DATA_BLOCK "DB_Scada_default"   // DB2112
{ S7_Optimized_Access := 'FALSE' }
VERSION : 0.1
   VAR
      tAlm : Struct   // HMI Alarms
         tE : Struct
            x0 : Bool;   // KE.Main emergency on
            x1 : Bool;   // KE1.Local emergency on
            x2 : Bool;   // Cabinet.Emergency localization
            x3 : Bool;   // SB1.Emergency localization
            x4 : Bool;   // SB2.Emergency localization
            x5 : Bool;
            x6 : Bool;
            x7 : Bool;
            x8 : Bool;
            x9 : Bool;
            x10 : Bool;
            x11 : Bool;
            x12 : Bool;
            x13 : Bool;
            x14 : Bool;
            x15 : Bool;
            x16 : Bool;
            x17 : Bool;
            x18 : Bool;
            x19 : Bool;
            x20 : Bool;
            x21 : Bool;
            x22 : Bool;
            x23 : Bool;
            x24 : Bool;
            x25 : Bool;
            x26 : Bool;
            x27 : Bool;
            x28 : Bool;
            x29 : Bool;
            x30 : Bool;
            x31 : Bool;
         END_STRUCT;
         tS : Struct
            tS0 : Struct
               x0 : Bool;
               x1 : Bool;   // Syncro.YCut meter gap outside the limits
               x2 : Bool;
               x3 : Bool;
               x4 : Bool;
               x5 : Bool;
               x6 : Bool;
               x7 : Bool;
               x8 : Bool;   // xB21QF1.Power supply 24V logic
               x9 : Bool;
               x10 : Bool;   // Syncro.Main line meter gap outside the limits
               x11 : Bool;
               x12 : Bool;
               x13 : Bool;
               x14 : Bool;
               x15 : Bool;
               x16 : Bool;
               x17 : Bool;
               x18 : Bool;
               x19 : Bool;
               x20 : Bool;
               x21 : Bool;
               x22 : Bool;
               x23 : Bool;
               x24 : Bool;
               x25 : Bool;
               x26 : Bool;
               x27 : Bool;
               x28 : Bool;
               x29 : Bool;
               x30 : Bool;
               x31 : Bool;
            END_STRUCT;
            tS1 : Struct
               x0 : Bool;
               x1 : Bool;   // Syncro.YCut meter gap outside the limits
               x2 : Bool;
               x3 : Bool;
               x4 : Bool;
               x5 : Bool;
               x6 : Bool;
               x7 : Bool;
               x8 : Bool;   // xB21QF1.Power supply 24V logic
               x9 : Bool;
               x10 : Bool;   // Syncro.Main line meter gap outside the limits
               x11 : Bool;
               x12 : Bool;
               x13 : Bool;
               x14 : Bool;
               x15 : Bool;
               x16 : Bool;
               x17 : Bool;
               x18 : Bool;
               x19 : Bool;
               x20 : Bool;
               x21 : Bool;
               x22 : Bool;
               x23 : Bool;
               x24 : Bool;
               x25 : Bool;
               x26 : Bool;
               x27 : Bool;
               x28 : Bool;
               x29 : Bool;
               x30 : Bool;
               x31 : Bool;
            END_STRUCT;
            tS2 : Struct
               x0 : Bool;
               x1 : Bool;   // Syncro.YCut meter gap outside the limits
               x2 : Bool;
               x3 : Bool;
               x4 : Bool;
               x5 : Bool;
               x6 : Bool;
               x7 : Bool;
               x8 : Bool;   // xB21QF1.Power supply 24V logic
               x9 : Bool;
               x10 : Bool;   // Syncro.Main line meter gap outside the limits
               x11 : Bool;
               x12 : Bool;
               x13 : Bool;
               x14 : Bool;
               x15 : Bool;
               x16 : Bool;
               x17 : Bool;
               x18 : Bool;
               x19 : Bool;
               x20 : Bool;
               x21 : Bool;
               x22 : Bool;
               x23 : Bool;
               x24 : Bool;
               x25 : Bool;
               x26 : Bool;
               x27 : Bool;
               x28 : Bool;
               x29 : Bool;
               x30 : Bool;
               x31 : Bool;
            END_STRUCT;
            tS3 : Struct
               x0 : Bool;
               x1 : Bool;   // Syncro.YCut meter gap outside the limits
               x2 : Bool;
               x3 : Bool;
               x4 : Bool;
               x5 : Bool;
               x6 : Bool;
               x7 : Bool;
               x8 : Bool;   // xB21QF1.Power supply 24V logic
               x9 : Bool;
               x10 : Bool;   // Syncro.Main line meter gap outside the limits
               x11 : Bool;
               x12 : Bool;
               x13 : Bool;
               x14 : Bool;
               x15 : Bool;
               x16 : Bool;
               x17 : Bool;
               x18 : Bool;
               x19 : Bool;
               x20 : Bool;
               x21 : Bool;
               x22 : Bool;
               x23 : Bool;
               x24 : Bool;
               x25 : Bool;
               x26 : Bool;
               x27 : Bool;
               x28 : Bool;
               x29 : Bool;
               x30 : Bool;
               x31 : Bool;
            END_STRUCT;
         END_STRUCT;
         tF : Struct
            x0 : Bool;
            x1 : Bool;
            x2 : Bool;
            x3 : Bool;
            x4 : Bool;
            x5 : Bool;
            x6 : Bool;
            x7 : Bool;
            x8 : Bool;
            x9 : Bool;
            x10 : Bool;
            x11 : Bool;
            x12 : Bool;
            x13 : Bool;
            x14 : Bool;
            x15 : Bool;
            x16 : Bool;
            x17 : Bool;
            x18 : Bool;
            x19 : Bool;
            x20 : Bool;
            x21 : Bool;
            x22 : Bool;
            x23 : Bool;
            x24 : Bool;
            x25 : Bool;
            x26 : Bool;
            x27 : Bool;
            x28 : Bool;
            x29 : Bool;
            x30 : Bool;
            x31 : Bool;
         END_STRUCT;
         tW : Struct
            x0 : Bool;   // PLCA.Timeout receiving consumed message
            x1 : Bool;   // PLCB.Timeout receiving consumed message
            x2 : Bool;   // PLCA.Mission packet lost
            x3 : Bool;   // PLCB.Mission packet lost
            x4 : Bool;   // PLCA.Syncro packet lost
            x5 : Bool;   // PLCB.Syncro packet lost
            x6 : Bool;   // QF.Protection air conditioners
            x7 : Bool;
            x8 : Bool;
            x9 : Bool;
            x10 : Bool;
            x11 : Bool;
            x12 : Bool;
            x13 : Bool;
            x14 : Bool;
            x15 : Bool;
            x16 : Bool;
            x17 : Bool;
            x18 : Bool;
            x19 : Bool;
            x20 : Bool;
            x21 : Bool;
            x22 : Bool;
            x23 : Bool;
            x24 : Bool;
            x25 : Bool;
            x26 : Bool;
            x27 : Bool;
            x28 : Bool;
            x29 : Bool;
            x30 : Bool;
            x31 : Bool;
         END_STRUCT;
      END_STRUCT;
      tHMR : Struct   // HMI Read
         xSpare0 : Bool := FALSE;   // Calibration function allowed {x|x|x|x|O}
         xSpare1 : Bool;
         xSpare2 : Bool;
         xSpare3 : Bool;
         xSpare4 : Bool;
         xSpare5 : Bool;
         xSpare6 : Bool;
         xSpare7 : Bool;
         xSpare8 : Bool;
         xSpare9 : Bool;
         xSpare10 : Bool;
         xSpare11 : Bool;
         xSpare12 : Bool;
         xSpare13 : Bool;
         xSpare14 : Bool;
         xSpare15 : Bool := FALSE;
         xSpare16 : Bool;
         xSpare17 : Bool;
         xSpare18 : Bool;
         xSpare19 : Bool;
         xSpare20 : Bool;
         xSpare21 : Bool;
         xSpare22 : Bool;
         xSpare23 : Bool;
         xSpare24 : Bool;
         xSpare25 : Bool;
         xSpare26 : Bool;
         xSpare27 : Bool;
         xSpare28 : Bool;
         xSpare29 : Bool;
         xSpare30 : Bool;
         xSpare31 : Bool;
         xSpare : Array[0..15] of Bool;
         iSpare0 : Int;
         iSpare1 : Int;
         iSpare2 : Int;
         iSpare3 : Int;
         iSpare4 : Int;
         iSpare5 : Int;
         iSpare6 : Int;
         iSpare7 : Int;
         iSpare8 : Int;
         iSpare9 : Int;
         iSpare10 : Int;
         iSpare11 : Int;
         iSpare12 : Int;
         iSpare13 : Int;
         iSpare14 : Int;
         iSpare15 : Int;
         iSpare16 : Int;
         dSpare0 : DInt := 0;   // Zone modality (1=Manual;4=Automatic;8=Manual request) {x|x|x|x|O}
         dSpare1 : DInt := 0;   // HMI Alarms
         dSpare2 : DInt := 0;   // HMI Write
         dSpare3 : DInt := 0;   // Production modality request (1=Out of Production 3= In production) {x|x|x|x|O}
         dSpare4 : DInt := 0;   // Production modality actual (1=Out of production 3=In production 8=Out of production request 9=In production request) {x|x|x|x|O}
         dSpare5 : DInt := 0;
         dSpare6 : DInt := 0;
         dSpare7 : DInt := 0;
         dSpare8 : DInt := 0;
         dSpare9 : DInt := 0;
         dSpare10 : DInt := 0;
         dSpare11 : DInt := 0;
         dSpare12 : DInt;
         dSpare13 : DInt;
         dSpare14 : DInt;
         dSpare15 : DInt;
         dSpare : Array[0..15] of DInt;
         rSpare0 : Real;
         rSpare1 : Real;
         rSpare2 : Real;
         rSpare3 : Real;
         rSpare4 : Real;
         rSpare5 : Real;
         rSpare6 : Real;
         rSpare7 : Real;
         rSpare8 : Real;
         tManCmd : Struct
            xSpare0 : Bool;
            xSpare1 : Bool;
            xSpare2 : Bool;
            xSpare3 : Bool;
            xSpare4 : Bool;
            xSpare5 : Bool;
            xSpare6 : Bool;
            xSpare7 : Bool;
            xSpare8 : Bool;
            xSpare9 : Bool;
            xSpare10 : Bool;
            xSpare11 : Bool;
            xSpare12 : Bool;
            xSpare13 : Bool;
            xSpare14 : Bool;
            xSpare15 : Bool;
            xSpare : Array[0..15] of Bool;
         END_STRUCT;
      END_STRUCT;
      tHMW : Struct   // HMI Write
         xSpare0 : Bool := FALSE;   // Automatic mode request {x|x|x|x|O}
         xSpare1 : Bool := FALSE;   // Manual mode request {x|x|x|x|O}
         xSpare2 : Bool := FALSE;   // Bridge out of production request {x|x|x|x|O}
         xSpare3 : Bool := FALSE;   // Bridge in production request {x|x|x|x|O}
         xSpare4 : Bool := FALSE;   // Cut during glass break {x|x|x|x|O}
         xSpare5 : Bool := FALSE;   // Motors and cards initialize {x|x|x|x|M}
         xSpare6 : Bool := FALSE;   // Force the homing of the heads {x|x|x|x|M}
         xSpare7 : Bool := FALSE;   // Position calibration request {x|x|x|x|M}
         xSpare8 : Bool := FALSE;   // Bridge offset calibration request {x|x|x|x|M}
         xSpare9 : Bool;
         xSpare10 : Bool;
         xSpare11 : Bool;
         xSpare12 : Bool;
         xSpare13 : Bool;
         xSpare14 : Bool := FALSE;
         xSpare15 : Bool := FALSE;
         xSpare16 : Bool := TRUE;
         xSpare17 : Bool := TRUE;
         xSpare18 : Bool := TRUE;
         xSpare19 : Bool := TRUE;
         xSpare20 : Bool := TRUE;
         xSpare21 : Bool := TRUE;
         xSpare22 : Bool := TRUE;
         xSpare23 : Bool := TRUE;
         xSpare24 : Bool;
         xSpare25 : Bool;
         xSpare26 : Bool;
         xSpare27 : Bool;
         xSpare28 : Bool;
         xSpare29 : Bool;
         xSpare30 : Bool;
         xSpare31 : Bool;
         xSpare : Array[0..15] of Bool;
         iSpare0 : Int;
         iSpare1 : Int;
         iSpare2 : Int;
         iSpare3 : Int;
         iSpare4 : Int;
         iSpare5 : Int;
         iSpare6 : Int;
         iSpare7 : Int;
         iSpare8 : Int;
         iSpare9 : Int;
         iSpare10 : Int;
         iSpare11 : Int;
         iSpare12 : Int;
         iSpare13 : Int;
         iSpare14 : Int;
         iSpare15 : Int;
         iSpare16 : Int := 0;
         dSpare0 : DInt := 0;   // Calibration. number of lite on calibration {x|x|1|8|M}
         dSpare1 : DInt := 0;   // Calibration. Move all the heads of this offset {mm/100|mm|-100|100|M}
         dSpare2 : DInt := 0;   // Pressure scaler during sample plate [%] {%|%|0|100|O}
         dSpare3 : DInt := 0;
         dSpare4 : DInt;
         dSpare5 : DInt;
         dSpare6 : DInt;
         dSpare7 : DInt;
         dSpare8 : DInt;
         dSpare9 : DInt;
         dSpare10 : DInt;
         dSpare11 : DInt;
         dSpare12 : DInt;
         dSpare13 : DInt;
         dSpare14 : DInt;
         dSpare15 : DInt;
         dSpare16 : DInt;
         dSpare17 : DInt;
         dSpare18 : DInt;
         dSpare19 : DInt;
         dSpare20 : DInt;
         dSpare21 : DInt;
         dSpare22 : DInt;
         dSpare23 : DInt;
         dSpare24 : DInt;
         dSpare25 : DInt;
         dSpare26 : DInt;
         dSpare27 : DInt;
         dSpare28 : DInt;
         dSpare29 : DInt;
         dSpare30 : DInt;
         dSpare31 : DInt;
         dSpare32 : DInt;
         dSpare33 : DInt;
         dSpare34 : DInt;
         dSpare35 : DInt;
         dSpare36 : DInt;
         dSpare37 : DInt;
         dSpare38 : DInt;
         dSpare39 : DInt;
         dSpare : Array[0..19] of DInt;
         rSpare0 : Real;
         rSpare1 : Real;
         rSpare2 : Real;
         rSpare3 : Real;
         rSpare4 : Real;
         rSpare5 : Real;
         rSpare6 : Real;
         rSpare7 : Real;
         rSpare8 : Real;
         tManCmd : Struct
            xSpare0 : Bool := FALSE;
            xSpare1 : Bool := FALSE;
            xSpare2 : Bool;
            xSpare3 : Bool;
            xSpare4 : Bool;
            xSpare5 : Bool;
            xSpare6 : Bool;
            xSpare7 : Bool;
            xSpare8 : Bool;
            xSpare9 : Bool;
            xSpare10 : Bool;
            xSpare11 : Bool;
            xSpare12 : Bool;
            xSpare13 : Bool;
            xSpare14 : Bool;
            xSpare15 : Bool;
            xSpare16 : Bool;
            xSpare17 : Bool;
            xSpare18 : Bool;
            xSpare19 : Bool;
            xSpare20 : Bool;
            xSpare21 : Bool;
            xSpare22 : Bool;
            xSpare23 : Bool;
            xSpare24 : Bool;
            xSpare25 : Bool;
            xSpare26 : Bool;
            xSpare27 : Bool;
            xSpare28 : Bool;
            xSpare29 : Bool;
            xSpare30 : Bool;
            xSpare31 : Bool;
         END_STRUCT;
      END_STRUCT;
   END_VAR
BEGIN
END_DATA_BLOCK

// folder: Communication

DATA_BLOCK "CM_Manager"   // DB1
{ S7_Optimized_Access := 'TRUE' }
VERSION : 0.1
BEGIN
END_DATA_BLOCK

DATA_BLOCK "CM_IDEV_FromMainLine"   // DB2
{ S7_Optimized_Access := 'TRUE' }
VERSION : 0.1
BEGIN
END_DATA_BLOCK

DATA_BLOCK "CM_IDEV_ToMainLine"   // DB3
{ S7_Optimized_Access := 'TRUE' }
VERSION : 0.1
BEGIN
END_DATA_BLOCK

DATA_BLOCK "CM_RECV_MissionData"   // DB4
{ S7_Optimized_Access := 'TRUE' }
VERSION : 0.1
BEGIN
END_DATA_BLOCK

DATA_BLOCK "CM_RECV_SyncroData"   // DB8
{ S7_Optimized_Access := 'TRUE' }
VERSION : 0.1
BEGIN
END_DATA_BLOCK

DATA_BLOCK "CM_BRCV_FromMainLine0"   // DB12
{ S7_Optimized_Access := 'TRUE' }
VERSION : 0.1
BEGIN
END_DATA_BLOCK

DATA_BLOCK "CM_BRCV_FromMainLine1"   // DB24
{ S7_Optimized_Access := 'TRUE' }
VERSION : 0.1
BEGIN
END_DATA_BLOCK

// folder: ILx2_Blocks

DATA_BLOCK "ILx2T_Parameter_Initialize_DB"   // DB10
{ S7_Optimized_Access := 'TRUE' }
VERSION : 1.1
// stored: InstanceOfName ILx2T_Parameter_Read_Write
"ILx2T_Parameter_Read_Write"
BEGIN
END_DATA_BLOCK

// folder: Subroutine

DATA_BLOCK "OB_Initialize"   // DB18
{ S7_Optimized_Access := 'TRUE' }
AUTHOR : Cigliutt
FAMILY : GP
VERSION : 1.0
// stored: InstanceOfName GP_OB_Initialize
"GP_OB_Initialize"
BEGIN
END_DATA_BLOCK

// folder: TaskErrors

DATA_BLOCK "RALRM_AUX_DB"   // DB59
{ S7_Optimized_Access := 'TRUE' }
VERSION : 0.1
   VAR RETAIN
      tAlm : Struct   // HMI Alarms
         tS : Struct   // Stopping faults
            xSpare_0 : Bool := FALSE;
            xSpare_1 : Bool := FALSE;
            xSpare_2 : Bool := FALSE;
            xSpare_3 : Bool := FALSE;
            xSpare_4 : Bool := FALSE;
            xSpare_5 : Bool := FALSE;
            xSpare_6 : Bool := FALSE;
            xSpare_7 : Bool := FALSE;
            xSpare_8 : Bool := FALSE;
            xSpare_9 : Bool := FALSE;
            xSpare_10 : Bool := FALSE;
            xSpare_11 : Bool := FALSE;
            xSpare_12 : Bool := FALSE;
            xSpare_13 : Bool := FALSE;
            xSpare_14 : Bool := FALSE;
            xSpare_15 : Bool := FALSE;
            xSpare_16 : Bool := FALSE;
            xSpare_17 : Bool := FALSE;
            xSpare_18 : Bool := FALSE;
            xSpare_19 : Bool := FALSE;
            xSpare_20 : Bool := FALSE;
            xSpare_21 : Bool := FALSE;
            xSpare_22 : Bool := FALSE;
            xSpare_23 : Bool := FALSE;
            xSpare_24 : Bool := FALSE;
            xSpare_25 : Bool := FALSE;
            xSpare_26 : Bool := FALSE;
            xSpare_27 : Bool := FALSE;
            xSpare_28 : Bool := FALSE;
            xSpare_29 : Bool := FALSE;
            xSpare_30 : Bool := FALSE;
            xSpare_31 : Bool := FALSE;
         END_STRUCT;
         tF : Struct   // Faults
            xDevice1 : Bool := FALSE;   // R13QF1.R13QF2.Power failure 230v auxiliary / Status device error.Device#1
            xDevice2 : Bool := FALSE;   // R18QF3.Power supply 24v logic / Status device error.Device#2
            xDevice3 : Bool := FALSE;   // R18QF4.Power supply 24v logic / Status device error.Device#3
            xDevice4 : Bool := FALSE;   // R18AP1.Redundancy 24v ok / Status device error.Device#4
            xDevice5 : Bool := FALSE;   // Status device error.Device#5
            xDevice6 : Bool := FALSE;   // Status device error.Device#6
            xDevice7 : Bool := FALSE;   // Status device error.Device#7
            xDevice8 : Bool := FALSE;   // Status device error.Device#8
            xDevice9 : Bool := FALSE;   // Status device error.Device#9
            xDevice10 : Bool := FALSE;   // Status device error.Device#10
            xSpare_10 : Bool := FALSE;
            xSpare_11 : Bool := FALSE;
            xSpare_12 : Bool;
            xSpare_13 : Bool;   // M250.R12KM1.Feedback rotation
            xSpare_14 : Bool;
            xSpare_15 : Bool;
            xSpare_16 : Bool;
            xSpare_17 : Bool;   // R204SP1.Compressed air presence cutting bridges
            xSpare_18 : Bool;
            xSpare_19 : Bool;
            xSpare_20 : Bool := FALSE;
            xSpare_21 : Bool := FALSE;
            xSpare_22 : Bool := FALSE;
            xSpare_23 : Bool := FALSE;
            xSpare_24 : Bool := FALSE;
            xSpare_25 : Bool := FALSE;
            xSpare_26 : Bool := FALSE;
            xSpare_27 : Bool := FALSE;
            xSpare_28 : Bool := FALSE;
            xSpare_29 : Bool := FALSE;
            xSpare_30 : Bool := FALSE;
            xSpare_31 : Bool := FALSE;
         END_STRUCT;
         tW : Struct   // Warnings
            xSpare_0 : Bool := FALSE;
            xSpare_1 : Bool := FALSE;
            xSpare_2 : Bool := FALSE;
            xSpare_3 : Bool := FALSE;
            xSpare_4 : Bool := FALSE;
            xSpare_5 : Bool := FALSE;
            xSpare_6 : Bool := FALSE;
            xSpare_7 : Bool := FALSE;
            xSpare_8 : Bool := FALSE;
            xSpare_9 : Bool := FALSE;
            xSpare_10 : Bool := FALSE;
            xSpare_11 : Bool := FALSE;
            xSpare_12 : Bool := FALSE;
            xSpare_13 : Bool := FALSE;
            xSpare_14 : Bool := FALSE;
            xSpare_15 : Bool := FALSE;
            xSpare_16 : Bool := FALSE;
            xSpare_17 : Bool := FALSE;
            xSpare_18 : Bool := FALSE;
            xSpare_19 : Bool := FALSE;
            xSpare_20 : Bool := FALSE;
            xSpare_21 : Bool := FALSE;
            xSpare_22 : Bool := FALSE;
            xSpare_23 : Bool := FALSE;
            xSpare_24 : Bool := FALSE;
            xSpare_25 : Bool := FALSE;
            xSpare_26 : Bool := FALSE;
            xSpare_27 : Bool := FALSE;
            xSpare_28 : Bool := FALSE;
            xSpare_29 : Bool := FALSE;
            xSpare_30 : Bool := FALSE;
            xSpare_31 : Bool := FALSE;
         END_STRUCT;
      END_STRUCT;
   END_VAR
BEGIN
END_DATA_BLOCK

// folder: (top level)

FUNCTION_BLOCK "M256_Manager"   // FB11, LAD
TITLE = #### HEAD MANAGER ####
{ S7_Optimized_Access := 'TRUE' }
VERSION : 0.1
   VAR_INPUT
      IN_tConnectionData : Array[0.."CONST_dNumberOfHeadsCycle"] of "UDT_MB_ConnData";   // IP and connection ID
   END_VAR
   VAR
      M256M_IDB : Array[0.."CONST_dNumberOfHeadsCycle"] of "M256M";
      M256F_IDB : Array[0.."CONST_dNumberOfHeadsCycle"] of "M256F";
      M256A_IDB : Array[0.."CONST_dNumberOfHeadsCycle"] of "M256A";
      M256A_ST_xAllHeadStoppingFaults : Bool;   // Cumulative Head in alarm
      M256F_ST_xAllHeadStoppingFaults : Bool;   // Cumulative Head in alarm
      M256M_ST_xAllHeadStoppingFaults : Bool;   // Cumulative Head in alarm
      M256M_ST_xAllHeadInitialized : Bool;
      M256M_ST_xAllHeadReferred : Bool;
      M256M_ST_xAllHeadPositioned : Bool;
      M256M_ST_xAllHeadIPLinked : Bool;
   END_VAR
   VAR_TEMP
      TMP_rgxHeadReferredSwitch : Array[0.."CONST_dNumberOfHeadsCycle"] of Bool;
      TMP_rgxHeadVirtualCollision : Array[0.."CONST_dNumberOfHeadsCycle"] of Bool;
      TMP_OS_XBrakeRelease : Bool;
      TMP_OS_XBrakeEngage : Bool;
      TMP_xHeadReferredSwicth : Bool;
      TMP_dIndex : DInt;
      TMP_dIndex2Nd : DInt;
      TMP_xDummy : Bool;
   END_VAR
BEGIN

REGION Network 1: #### COSTANTS ####
END_REGION

REGION Network 2: #### ALARMS ####
END_REGION

REGION Network 3: Op. side head overstroke
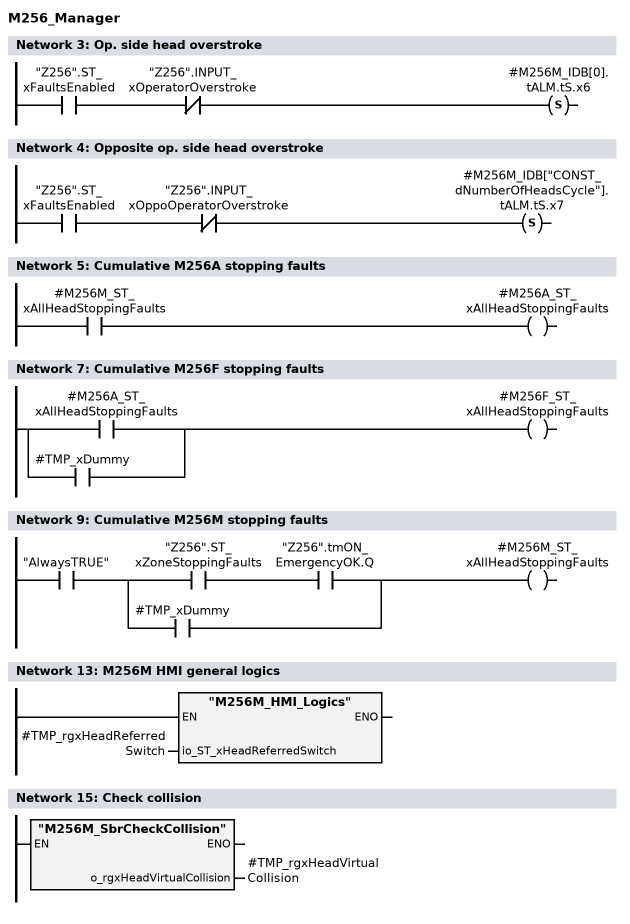
   RUNG wire#powerrail
      Contact( "Z256".ST_xFaultsEnabled )
      I_Contact( "Z256".INPUT_xOperatorOverstroke )
      S_Coil( #M256M_IDB[0].tALM.tS.x6 )
   END_RUNG
   // the same network as SCL:
   IF "Z256".ST_xFaultsEnabled AND NOT "Z256".INPUT_xOperatorOverstroke THEN
       #M256M_IDB[0].tALM.tS.x6 := TRUE;
   END_IF;
END_REGION

REGION Network 4: Opposite op. side head overstroke
   RUNG wire#powerrail
      Contact( "Z256".ST_xFaultsEnabled )
      I_Contact( "Z256".INPUT_xOppoOperatorOverstroke )
      S_Coil( #M256M_IDB["CONST_dNumberOfHeadsCycle"].tALM.tS.x7 )
   END_RUNG
   // the same network as SCL:
   IF "Z256".ST_xFaultsEnabled AND NOT "Z256".INPUT_xOppoOperatorOverstroke THEN
       #M256M_IDB["CONST_dNumberOfHeadsCycle"].tALM.tS.x7 := TRUE;
   END_IF;
END_REGION

REGION Network 5: Cumulative M256A stopping faults
   RUNG wire#powerrail
      Contact( #M256M_ST_xAllHeadStoppingFaults )
      Coil( #M256A_ST_xAllHeadStoppingFaults )
   END_RUNG
   // the same network as SCL:
   #M256A_ST_xAllHeadStoppingFaults := #M256M_ST_xAllHeadStoppingFaults;
END_REGION

REGION Network 6 (SCL): Cumulative M256F faults status
   #TMP_xDummy := FALSE;
   FOR #TMP_dIndex := 0 TO "CONST_dNumberOfHeadsCycle" DO
       IF #M256F_IDB[#TMP_dIndex].ST_xStoppingFaults THEN
           #TMP_xDummy := TRUE;
       END_IF;
   END_FOR;
END_REGION

REGION Network 7: Cumulative M256F stopping faults
   RUNG wire#powerrail
      Contact( #M256A_ST_xAllHeadStoppingFaults )
      wire#w1
      Coil( #M256F_ST_xAllHeadStoppingFaults )
   END_RUNG
   RUNG wire#powerrail
      Contact( #TMP_xDummy )
   END_RUNG wire#w1
   // the same network as SCL:
   #M256F_ST_xAllHeadStoppingFaults := #M256A_ST_xAllHeadStoppingFaults OR #TMP_xDummy;
END_REGION

REGION Network 8 (SCL): Cumulative M256M faults status
   #TMP_xDummy := FALSE;
   FOR #TMP_dIndex := 0 TO "CONST_dNumberOfHeadsCycle" DO
       IF #M256M_IDB[#TMP_dIndex].ST_xStoppingFaults THEN
           #TMP_xDummy := TRUE;
       END_IF;
   END_FOR;
END_REGION

REGION Network 9: Cumulative M256M stopping faults
   RUNG wire#powerrail
      Contact( "AlwaysTRUE" )
      wire#w1
      Contact( "Z256".ST_xZoneStoppingFaults )
      Contact( "Z256".tmON_EmergencyOK.Q )
      wire#w2
      Coil( #M256M_ST_xAllHeadStoppingFaults )
   END_RUNG
   RUNG wire#w1
      Contact( #TMP_xDummy )
   END_RUNG wire#w2
   // the same network as SCL:
   #M256M_ST_xAllHeadStoppingFaults := "AlwaysTRUE" AND (("Z256".ST_xZoneStoppingFaults AND "Z256".tmON_EmergencyOK.Q) OR #TMP_xDummy);
END_REGION

REGION Network 10: #### PHASES & LOGICS ####
END_REGION

REGION Network 11: #### M256M ####
END_REGION

REGION Network 12 (SCL): Compile data for Head referred array
   FOR #TMP_dIndex := 0 TO "CONST_dNumberOfHeadsCycle" DO
       #TMP_rgxHeadReferredSwitch[#TMP_dIndex] := #M256M_IDB[#TMP_dIndex].ST_xHeadReferredSwitch;
   END_FOR;
END_REGION

REGION Network 13: M256M HMI general logics
   RUNG wire#powerrail
      "M256M_HMI_Logics"(io_ST_xHeadReferredSwitch := #TMP_rgxHeadReferredSwitch)
   END_RUNG
   // the same network as SCL:
   "M256M_HMI_Logics"(io_ST_xHeadReferredSwitch := #TMP_rgxHeadReferredSwitch);
END_REGION

REGION Network 14 (SCL): Recompile data for Head referred array
   FOR #TMP_dIndex := 0 TO "CONST_dNumberOfHeadsCycle" DO
       #M256M_IDB[#TMP_dIndex].ST_xHeadReferredSwitch := #TMP_rgxHeadReferredSwitch[#TMP_dIndex];
   END_FOR;
END_REGION

REGION Network 15: Check collision
   RUNG wire#powerrail
      "M256M_SbrCheckCollision"(o_rgxHeadVirtualCollision => #TMP_rgxHeadVirtualCollision)
   END_RUNG
   // the same network as SCL:
   "M256M_SbrCheckCollision"(o_rgxHeadVirtualCollision => #TMP_rgxHeadVirtualCollision);
END_REGION

REGION Network 16 (SCL): Check head initialized, positioned, referred, communication
   #M256M_ST_xAllHeadInitialized := TRUE;
   #M256M_ST_xAllHeadReferred := TRUE;
   #M256M_ST_xAllHeadPositioned := TRUE;
   #M256M_ST_xAllHeadIPLinked := TRUE;


   //IF one head of the heads isn't TRUE reset "All head xxx" bit
   FOR #TMP_dIndex := 0 TO "CONST_dNumberOfHeadsCycle" DO
       IF NOT #M256M_IDB[#TMP_dIndex].ST_xHeadInitialized THEN
           #M256M_ST_xAllHeadInitialized := FALSE;
       END_IF;
       IF NOT #M256M_IDB[#TMP_dIndex].ST_xHeadPositioned THEN
           #M256M_ST_xAllHeadPositioned := FALSE;
       END_IF;
       IF NOT #M256M_IDB[#TMP_dIndex].ST_xHeadReferredSwitch THEN
           #M256M_ST_xAllHeadReferred := FALSE;
       END_IF;
       IF NOT #M256M_IDB[#TMP_dIndex].ST_xHeadIPAvail THEN
           #M256M_ST_xAllHeadReferred := FALSE;
       END_IF;
   END_FOR;
END_REGION

REGION Network 17 (SCL): Call M256M logic

   FOR #TMP_dIndex := 0 TO "CONST_dNumberOfHeadsCycle" DO

       //Compile data for FB
       #M256M_IDB[#TMP_dIndex].ST_xHeadVirtualCollision := #TMP_rgxHeadVirtualCollision[#TMP_dIndex];
       //Call Move manager
       #M256M_IDB[#TMP_dIndex](IN_dHeadCycleIndex := #TMP_dIndex,
                                   IN_tConnectionData := #IN_tConnectionData[#TMP_dIndex],
                                   IN_ST_xAllHeadInitialized := #M256M_ST_xAllHeadInitialized,
                                   IN_ST_xAllHeadReferred := #M256M_ST_xAllHeadReferred,
                                   IN_ST_xAllHeadPositioned := #M256M_ST_xAllHeadPositioned,
                                   IN_xST_AllHeadStoppingFaults:= #M256M_ST_xAllHeadStoppingFaults);

   END_FOR;
END_REGION

REGION Network 18 (SCL): Move cadencer
   //   Description: This function will cadencer the movement to avoid collision problem

   FOR #TMP_dIndex := 0 TO "CONST_dNumberOfHeadsCycle" DO

       //Check if the movement is request for the head
       IF #M256M_IDB[#TMP_dIndex].PH_xHeadPositioning AND #M256A_IDB[#TMP_dIndex].ST_xCarriageUpPosition THEN

           //If to home let the movement
           IF #M256M_IDB[#TMP_dIndex].AUX_dHeadRequestPosition_cmm = #M256M_IDB[#TMP_dIndex].tHMR.dHeadHomePositions_cmm THEN
               #M256M_IDB[#TMP_dIndex].AUX_xPosCadencer := TRUE;
           END_IF;

           //Ok. Movement is requested. Check if is request a operator movement or opposite operator movement
           IF #M256M_IDB[#TMP_dIndex].AUX_dHeadRequestPosition_cmm >= #M256M_IDB[#TMP_dIndex].AUX_dHeadActualPosition_cmm THEN

               //Is requested an to opposite operator movement. Check the state of the next head.
               //The condition to allow the movement are:
               //1. Is the last head
               //2. The target position is less then the actual position of the next head.
               //3. The target position is more then the actual position of the next head, but the next head has the feedback of movement in progress
               IF #TMP_dIndex = ("CONST_dNumberOfHeads" - 1) THEN
                   #M256M_IDB[#TMP_dIndex].AUX_xPosCadencer := TRUE;
               ELSIF ((#M256M_IDB[#TMP_dIndex].AUX_dHeadRequestPosition_cmm + "PLANT_CONSTANTS".CONST_dHOppoSideEnc_cmm[#TMP_dIndex]) <
                   (#M256M_IDB[#TMP_dIndex + 1].AUX_dHeadActualPosition_cmm - "PLANT_CONSTANTS".CONST_dHOpSideEnc_cmm[#TMP_dIndex + 1])) THEN
                   #M256M_IDB[#TMP_dIndex].AUX_xPosCadencer := TRUE;
               ELSIF #M256M_IDB[#TMP_dIndex + 1].ST_xMovementInProgress THEN
                   #M256M_IDB[#TMP_dIndex].AUX_xPosCadencer := TRUE;
               END_IF;

           ELSE

               //Is requested an to operator movement. Check the state of the previous head.
               //The condition to allow the movement are:
               //1. Is the first head
               //2. The target position is greather then the actual position of the previous head.
               //3. The target position is less then the actual position of the previous head, but the previous head has the feedback of movement in progress
               IF (#TMP_dIndex = 0) THEN
                   #M256M_IDB[#TMP_dIndex].AUX_xPosCadencer := 1;
               ELSIF ((#M256M_IDB[#TMP_dIndex].AUX_dHeadRequestPosition_cmm - "PLANT_CONSTANTS".CONST_dHOpSideEnc_cmm[#TMP_dIndex]) >
                   (#M256M_IDB[#TMP_dIndex - 1].AUX_dHeadActualPosition_cmm + "PLANT_CONSTANTS".CONST_dHOppoSideEnc_cmm[#TMP_dIndex - 1])) THEN
                   #M256M_IDB[#TMP_dIndex].AUX_xPosCadencer := 1;
               ELSIF #M256M_IDB[#TMP_dIndex -1].ST_xMovementInProgress THEN

                   #M256M_IDB[#TMP_dIndex].AUX_xPosCadencer := 1;
               END_IF;
           END_IF;
       END_IF;


       //Check if the movement is request for the head
       IF #M256M_IDB[#TMP_dIndex].PH_xHeadHomeSwitch THEN

           //Check the home direction of the head. 
           IF NOT "PLANT_CONSTANTS".CONST_rgxHomeSide[#TMP_dIndex] THEN

               //Head direction to operator side. The condition to allow the movement are
               //1. Is the first head
               //2. The previous head already home
               //3. The previous head already start the home
               IF #TMP_dIndex = 0 THEN
                   #M256M_IDB[#TMP_dIndex].AUX_xHomeCadencer := TRUE;
               ELSIF #M256M_IDB[#TMP_dIndex - 1].ST_xHeadReferredSwitch THEN
                   #M256M_IDB[#TMP_dIndex].AUX_xHomeCadencer := TRUE;
               ELSIF #M256M_IDB[#TMP_dIndex - 1].ILx2T_Homing_Instance.q_xBusy THEN
                   #M256M_IDB[#TMP_dIndex].AUX_xHomeCadencer := TRUE;
               END_IF;
           ELSE
               //Head direction to opposite operator side. The condition to allow the movement are
               //1. Is the last head
               //2. The previous head already home
               //3. The previous head already start the home
               IF #TMP_dIndex = "CONST_dNumberOfHeads" - 1 THEN
                   #M256M_IDB[#TMP_dIndex].AUX_xHomeCadencer := TRUE;
               ELSIF #M256M_IDB[#TMP_dIndex + 1].ST_xHeadReferredSwitch THEN
                   #M256M_IDB[#TMP_dIndex].AUX_xHomeCadencer := TRUE;
               ELSIF #M256M_IDB[#TMP_dIndex + 1].ILx2T_Homing_Instance.q_xBusy THEN
                   #M256M_IDB[#TMP_dIndex].AUX_xHomeCadencer := TRUE;
               END_IF;
           END_IF;
       END_IF;
   END_FOR;
END_REGION

REGION Network 19: #### M256A ####
END_REGION

REGION Network 20 (SCL): Move mission manager
   FOR #TMP_dIndex := 0 TO "CONST_dNumberOfHeadsCycle" DO

       //Check the request. If rise allow without control.
       //If descent check if the position of the ycut is matching the request position.
       IF "Z256_Manager".tOutputData.rgxArmRequest[#TMP_dIndex] AND #M256M_IDB[#TMP_dIndex].IN_ST_xAllHeadPositioned AND
           (#M256M_IDB[#TMP_dIndex].AUX_dHeadRequestPosition_cmm = "Z256_Manager".tOutputData.rgdHeadsPositions_cmm[#TMP_dIndex]) THEN
           #M256A_IDB[#TMP_dIndex].AUX_xHeadArmRequest := 1;
       ELSE
           #M256A_IDB[#TMP_dIndex].AUX_xHeadArmRequest := 0;
       END_IF;

   END_FOR;
END_REGION

REGION Network 21 (SCL): Call M256A logics
   FOR #TMP_dIndex := 0 TO "CONST_dNumberOfHeadsCycle" DO
       #TMP_xDummy := false;
           IF NOT #M256M_IDB[#TMP_dIndex].ILx2T_Control_Instance.q_xSwitchedOn OR #M256M_ST_xAllHeadPositioned THEN
               #TMP_xDummy := true;
           END_IF;
           #M256A_IDB[#TMP_dIndex](IN_dHeadCycleIndex := #TMP_dIndex,
                                       IN_xDriveDisabled := #TMP_xDummy,
                                      IN_xST_AllHeadStoppingFaults := #M256A_ST_xAllHeadStoppingFaults);
   END_FOR;
END_REGION

REGION Network 22: #### M256F ####
END_REGION

REGION Network 23 (SCL): Call M256F logics
   FOR #TMP_dIndex := 0 TO "CONST_dNumberOfHeadsCycle" DO
       #M256F_IDB[#TMP_dIndex](IN_dHeadCycleIndex := #TMP_dIndex,
                                       IN_xHeadDescent := #M256A_IDB[#TMP_dIndex].OUTPUT_xCarriageDescent,
                                       IN_xST_AllHeadStoppingFaults := #M256F_ST_xAllHeadStoppingFaults);
   END_FOR;
END_REGION
END_FUNCTION_BLOCK

FUNCTION_BLOCK "M256A"   // FB12, LAD
{ S7_Optimized_Access := 'TRUE' }
VERSION : 0.1
   VAR_INPUT
      IN_xDriveDisabled : Bool;   // M256M drive disabled
      IN_dHeadCycleIndex : DInt;   // Number of head cycle (Actual head-1)
      IN_xST_AllHeadStoppingFaults : Bool;   // Cumulative head alarm
   END_VAR
   VAR
      ST_xOutputEnable : Bool;   // Head #x output enable
      ST_xPhaseInProgress : Bool;   // Head #x phases in progress
      ST_xWarnings : Bool;   // Head #x in warning
      ST_xFaults : Bool;   // Head #x in faults
      ST_xStoppingFaults : Bool;   // Head #x in stopping fault
      ST_xCarriageUpPosition : Bool;   // Status carriage head#x up position
      ST_xCarriageDownPosition : Bool;   // Status carriage head#x down position
      PH_xCarriageDescent : Bool;   // Head#x carriage descent in progress
      PH_xEndCarriageDescent : Bool;   // Head#x end carriage descent in progress
      PH_xCarriageRise : Bool;   // Head#x carriage rise in progress
      PH_xEndCarriageRise : Bool;   // Head#x end carriage rise in progress
      AUX_xHeadArmRequest : Bool;   // Head#x arm request from manager
      AUX_tmON_HeadDescent : IEC_TIMER;   // Head#x timer head descent
      AUX_tmON_HeadRise : IEC_TIMER;   // Head#x timer head rise
      AUX_tmON_FaultsCarrPos : IEC_TIMER;   // Head#x timer delay carriage in position
      AUX_tmOFF_FaultsCarrPos : IEC_TIMER;   // Head#x timer retain carriage in position
      INPUT_xForceArming : Bool;   // Head #x force arming
      INPUT_xHeadsUpIstan : Bool;   // Heads up istantaneous button
      INPUT_xCarriageInWorkPosition : Bool;   // Head#x carriage in work position
      OUTPUT_xCarriageDescent : Bool;   // Head#x carriage descent
      tALM : Struct
         tW : Struct
            x0 : Bool;
            x1 : Bool;
            x2 : Bool;
            x3 : Bool;
            x4 : Bool;
            x5 : Bool;
            x6 : Bool;
            x7 : Bool;
            x8 : Bool;
            x9 : Bool;
            x10 : Bool;
            x11 : Bool;
            x12 : Bool;
            x13 : Bool;
            x14 : Bool;
            x15 : Bool;
            x16 : Bool;
            x17 : Bool;
            x18 : Bool;
            x19 : Bool;
            x20 : Bool;
            x21 : Bool;
            x22 : Bool;
            x23 : Bool;
            x24 : Bool;
            x25 : Bool;
            x26 : Bool;
            x27 : Bool;
            x28 : Bool;
            x29 : Bool;
            x30 : Bool;
            x31 : Bool;
         END_STRUCT;
         tS : Struct
            xNotWorkPos : Bool;   // Head#x carriage not in working position
            x1 : Bool;
            x2 : Bool;
            x3 : Bool;
            x4 : Bool;
            x5 : Bool;
            x6 : Bool;
            x7 : Bool;
            x8 : Bool;
            x9 : Bool;
            x10 : Bool;
            x11 : Bool;
            x12 : Bool;
            x13 : Bool;
            x14 : Bool;
            x15 : Bool;
            x16 : Bool;
            x17 : Bool;
            x18 : Bool;
            x19 : Bool;
            x20 : Bool;
            x21 : Bool;
            x22 : Bool;
            x23 : Bool;
            x24 : Bool;
            x25 : Bool;
            x26 : Bool;
            x27 : Bool;
            x28 : Bool;
            x29 : Bool;
            x30 : Bool;
            x31 : Bool;
         END_STRUCT;
         tF : Struct
            x0 : Bool;
            x1 : Bool;
            x2 : Bool;
            x3 : Bool;
            x4 : Bool;
            x5 : Bool;
            x6 : Bool;
            x7 : Bool;
            x8 : Bool;
            x9 : Bool;
            x10 : Bool;
            x11 : Bool;
            x12 : Bool;
            x13 : Bool;
            x14 : Bool;
            x15 : Bool;
            x16 : Bool;
            x17 : Bool;
            x18 : Bool;
            x19 : Bool;
            x20 : Bool;
            x21 : Bool;
            x22 : Bool;
            x23 : Bool;
            x24 : Bool;
            x25 : Bool;
            x26 : Bool;
            x27 : Bool;
            x28 : Bool;
            x29 : Bool;
            x30 : Bool;
            x31 : Bool;
         END_STRUCT;
      END_STRUCT;
   END_VAR
   VAR RETAIN
      tHMR : Struct   // {[Unit][Scada unit][Low limit][High limit][Access]}
         dHeadStatus : DInt;   // Head#x arming status (1=Up 3=Down 7=Anomaly) {x|x|x|x|O}
         tManCmd : Struct
            xMan_DescentFdbk : Bool;   // Head #x manual descent feedback {x|x|x|x|O}
            xMan_RiseFdbk : Bool;   // Head #x manual rise feedback {x|x|x|x|O}
         END_STRUCT;
      END_STRUCT;
      tHMW : Struct   // {[Unit][Scada unit][Low limit][High limit][Access]}
         dRaiseReactTime_ms : DInt;   // Head#x raise reaction time [ms] {ms|s|-200|200|M}
         dDescentReactTime_ms : DInt;   // Head#x descent reaction time [ms] {ms|s|0|3000|M}
         tManCmd : Struct
            xManDescent : Bool;   // Head #x manual Descent {x|x|x|x|O}
            xManRise : Bool;   // Head #x manual rise {x|x|x|x|O}
         END_STRUCT;
      END_STRUCT;
   END_VAR
   VAR_TEMP
      TMP_dwDummy : DWord;
   END_VAR
   VAR_TEMP   // added for the SCL form of the ladder/FBD networks
      _w1 : Bool;
   END_VAR
BEGIN

REGION Network 1: ####_COSTANTS_####
END_REGION

REGION Network 2: ####_ALARMS_####
END_REGION

REGION Network 3: Reset faults